(* Logix 5000 project; controller PLC_MCC1201_220AP1 vendor 1 type 14 code 164 rev 35.11; software revision 35.00; part 20 of 25 *)
(* tags used below, declared in another part *)
   LEHR_dActualSpeedValue_mm_min : DINT;
   LEHR_dActualSpeedValueToConveyor_mm_min : DINT;
   LEHR_dLehrPositionAdvancement : DINT;
   SnaprollUPS_DistanceFromSnaproll_cmm : DINT;
   SnaprollUPS_xOS_NewCut : BOOL;
   SnaprollUPS_xOSR : BOOL;
   SnaprollUPS_xOutputRise : BOOL;
   tmOF_retainSnaprolUPS : TIMER;
   TMP_dDummy : DINT;
   TMP_dEncoderCutPosition : DINT;
   TMP_xCutOnSnaproll_cmm : BOOL;
   B3 : DINT[102];
   DISTANCE : ALIAS FOR N7[1];
   M203DROP : MAC_DROPCONV;
   M203DROP_ALM : MAC_DROPCONV_ALM;
   M203DROP_HMR : MAC_DROPCONV_HMR;
   M203DROP_HMW : MAC_DROPCONV_HMW;
   M225 : MAC_EMERGENCYXCUT;
   O : INT[128];
   Status : INT;   // INT tag to retrieve Status value through GSV created during conversion
   TMP_xAlwaysOFF : BOOL;
   TMP_xTestCycle : BOOL;
   W_APC_ACTIVE : ALIAS FOR W_B3[0].10;
   W_APC_BUTTON : ALIAS FOR W_I[8].10;
   W_B3 : DINT[7];
   W_BLOWDOWN_VALVE : ALIAS FOR W_O[10].12;
   W_CB1_START : ALIAS FOR W_O[10].1;
   W_CB2_START : ALIAS FOR W_O[10].3;
   W_COMPUTE_TCD3 : ALIAS FOR W_N7[923];
   W_COMPUTE_TCD5B : ALIAS FOR W_N7[926];
   W_CONDUCT_SENSOR : ALIAS FOR W_N7[110];
   W_CONV_PID_N7_620 : PID;   // Return Water Flow Control Valve Position
   W_CONV_PID_N7_650 : PID;   // RO Unit Water Temperature Control
   W_CONV_PID_N7_680 : PID;   // Boiler Water Temperature Control
   W_CONV_PID_N7_710 : PID;   // Mixed Air Control Damper Positioning
   W_CONV_PID_N7_740 : PID;   // Dryer Room Temperature Control
   W_CP1_ENABLE : ALIAS FOR W_B3[0].5;
   W_CP1A_START : ALIAS FOR W_O[10].5;
   W_CP1B_START : ALIAS FOR W_O[10].7;
   W_CP2A_START : ALIAS FOR W_O[10].9;
   W_CP2B_START : ALIAS FOR W_O[10].11;
   W_DRYER_PID_OUT : ALIAS FOR W_N7[925];
   W_EMER_STOP : ALIAS FOR W_I[8].13;
   W_FLOW_ENABLE : ALIAS FOR W_B3[0].9;
   W_HX1_BCD_OUT : ALIAS FOR W_N7[917];
   W_HX2_SENSOR : ALIAS FOR W_N7[47];
   W_I : INT[32];
   W_MA_FAN_SENSOR : ALIAS FOR W_N7[50];
   W_N11 : DINT[10];
   W_N7 : DINT[933];
   W_PID_INT_TO_TOD : ALIAS FOR W_N7[919];
   W_PS1_SWITCH : ALIAS FOR W_I[8].8;
   W_PWT_HIGH_LIMIT : ALIAS FOR W_I[8].2;
   W_RECIEVING_LEVEL : ALIAS FOR W_I[8].9;
   W_RET_PID_OUTPUT : ALIAS FOR W_N7[921];
   W_RO_START : ALIAS FOR W_O[10].13;
   W_RUN_WASHER : ALIAS FOR W_B3[0].2;
   W_SHUTDOWN_LATCH : ALIAS FOR W_B3[0].1;
   W_T4 : TIMER[101];
   W_TCD3_OUTPUT : ALIAS FOR W_N7[300];
   W_TCD3_PID_OUTPUT : ALIAS FOR W_N7[922];
   W_TCD4_OUTPUT : ALIAS FOR W_N7[301];
   W_TCD5A_OUTPUT : ALIAS FOR W_N7[302];
   W_TT3_RAW_BCD : ALIAS FOR W_N7[48];
   W_TT6_HITEMP_AIR : ALIAS FOR W_N7[49];
   Z200_UPS : ZONE_UPS;
(* MainProgram, continued *)

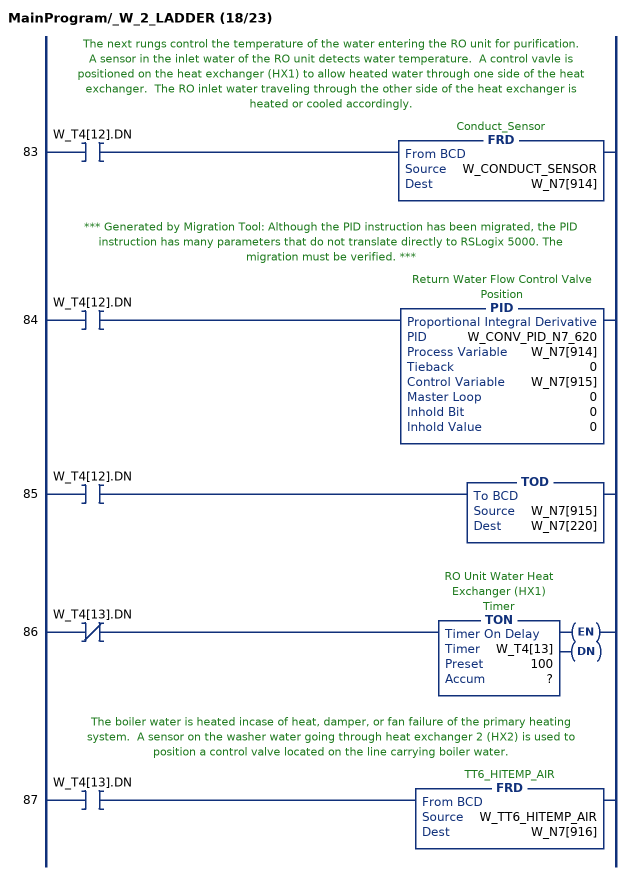
   [picture p330: MainProgram/_W_2_LADDER rungs 83-87]
   // The next rungs control the temperature of the water entering the RO unit for purification.  A sensor in the inlet water of the RO unit detects water temperature.  A control vavle is positioned on the heat exchanger (HX1) to allow heated water through one side of the heat exchanger.  The RO inlet water traveling through the other side of the heat exchanger is heated or cooled accordingly.
   83: XIC(W_T4[12].DN)FRD(W_CONDUCT_SENSOR,W_N7[914]);
   // *** Generated by Migration Tool: Although the PID instruction has been migrated, the PID instruction has many parameters that do not translate directly to RSLogix 5000. The migration must be verified. ***
   84: XIC(W_T4[12].DN)PID(W_CONV_PID_N7_620,W_N7[914],0,W_N7[915],0,0,0);
   85: XIC(W_T4[12].DN)TOD(W_N7[915],W_N7[220]);
   86: XIO(W_T4[13].DN)TON(W_T4[13],?,?);
   // The boiler water is heated incase of heat, damper, or fan failure of the primary heating system.  A sensor on the washer water going through heat exchanger 2 (HX2) is used to position a control valve located on the line carrying boiler water.
   87: XIC(W_T4[13].DN)FRD(W_TT6_HITEMP_AIR,W_N7[916]);
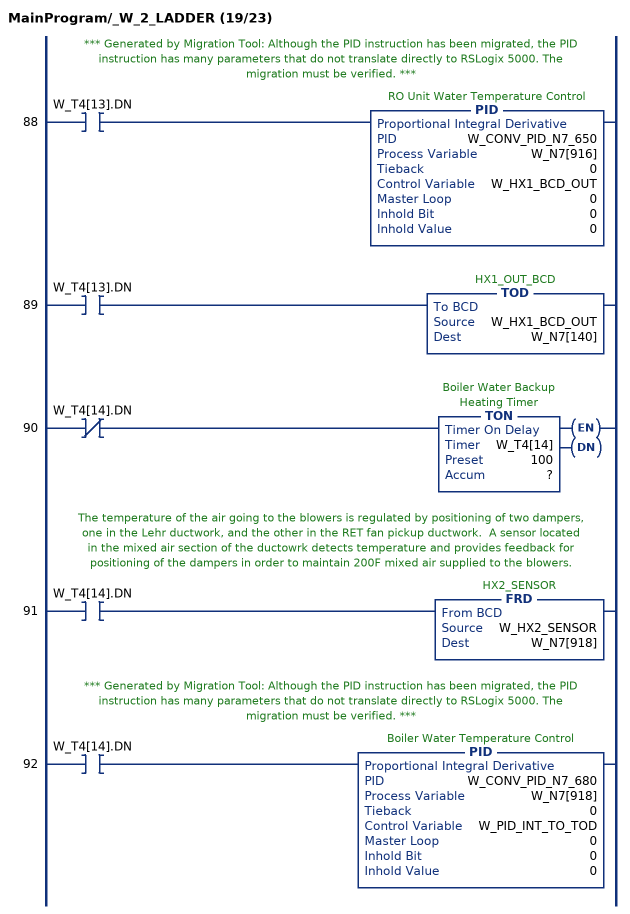
   // *** Generated by Migration Tool: Although the PID instruction has been migrated, the PID instruction has many parameters that do not translate directly to RSLogix 5000. The migration must be verified. ***
   88: XIC(W_T4[13].DN)PID(W_CONV_PID_N7_650,W_N7[916],0,W_HX1_BCD_OUT,0,0,0);
   89: XIC(W_T4[13].DN)TOD(W_HX1_BCD_OUT,W_N7[140]);
   90: XIO(W_T4[14].DN)TON(W_T4[14],?,?);
   // The temperature of the air going to the blowers is regulated by positioning of two dampers, one in the Lehr ductwork, and the other in the RET fan pickup ductwork.  A sensor located in the mixed air section of the ductowrk detects temperature and provides feedback for positioning of the dampers in order to maintain 200F mixed air supplied to the blowers.
   91: XIC(W_T4[14].DN)FRD(W_HX2_SENSOR,W_N7[918]);
   // *** Generated by Migration Tool: Although the PID instruction has been migrated, the PID instruction has many parameters that do not translate directly to RSLogix 5000. The migration must be verified. ***
   92: XIC(W_T4[14].DN)PID(W_CONV_PID_N7_680,W_N7[918],0,W_PID_INT_TO_TOD,0,0,0);
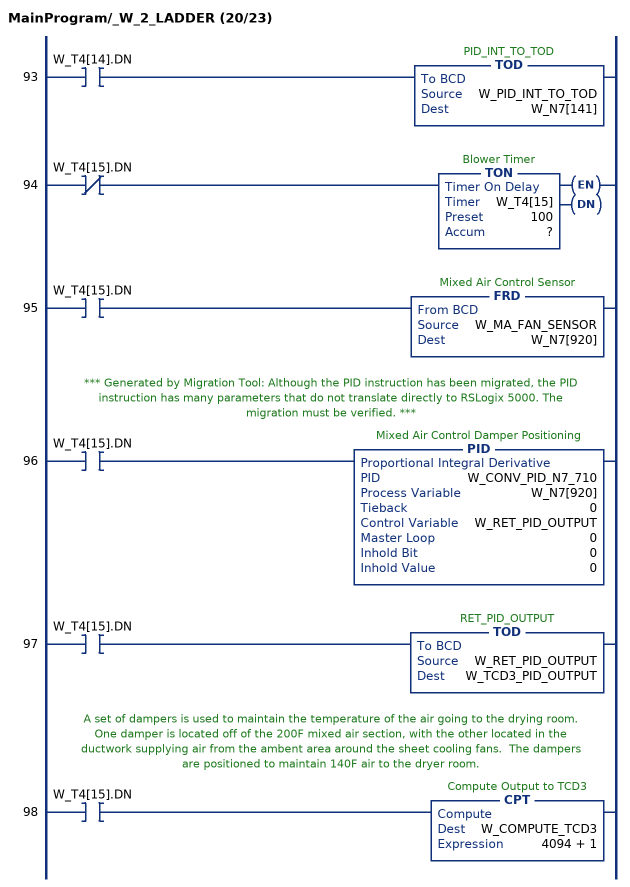
   93: XIC(W_T4[14].DN)TOD(W_PID_INT_TO_TOD,W_N7[141]);
   94: XIO(W_T4[15].DN)TON(W_T4[15],?,?);
   95: XIC(W_T4[15].DN)FRD(W_MA_FAN_SENSOR,W_N7[920]);
   // *** Generated by Migration Tool: Although the PID instruction has been migrated, the PID instruction has many parameters that do not translate directly to RSLogix 5000. The migration must be verified. ***
   96: XIC(W_T4[15].DN)PID(W_CONV_PID_N7_710,W_N7[920],0,W_RET_PID_OUTPUT,0,0,0);
   97: XIC(W_T4[15].DN)TOD(W_RET_PID_OUTPUT,W_TCD3_PID_OUTPUT);
   // A set of dampers is used to maintain the temperature of the air going to the drying room.  One damper is located off of the 200F mixed air section, with the other located in the ductwork supplying air from the ambent area around the sheet cooling fans.  The dampers are positioned to maintain 140F air to the dryer room.
   98: XIC(W_T4[15].DN)CPT(W_COMPUTE_TCD3,4094 + 1);
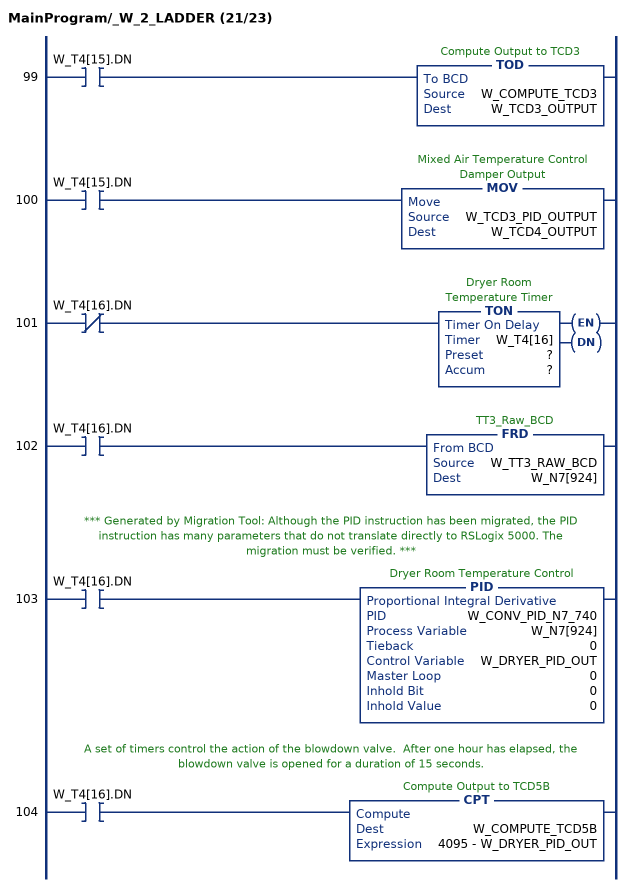
   99: XIC(W_T4[15].DN)TOD(W_COMPUTE_TCD3,W_TCD3_OUTPUT);
   100: XIC(W_T4[15].DN)MOV(W_TCD3_PID_OUTPUT,W_TCD4_OUTPUT);
   101: XIO(W_T4[16].DN)TON(W_T4[16],?,?);
   102: XIC(W_T4[16].DN)FRD(W_TT3_RAW_BCD,W_N7[924]);
   // *** Generated by Migration Tool: Although the PID instruction has been migrated, the PID instruction has many parameters that do not translate directly to RSLogix 5000. The migration must be verified. ***
   103: XIC(W_T4[16].DN)PID(W_CONV_PID_N7_740,W_N7[924],0,W_DRYER_PID_OUT,0,0,0);
   // A set of timers control the action of the blowdown valve.  After one hour has elapsed, the blowdown valve is opened for a duration of 15 seconds.
   104: XIC(W_T4[16].DN)CPT(W_COMPUTE_TCD5B,4095 - W_DRYER_PID_OUT);
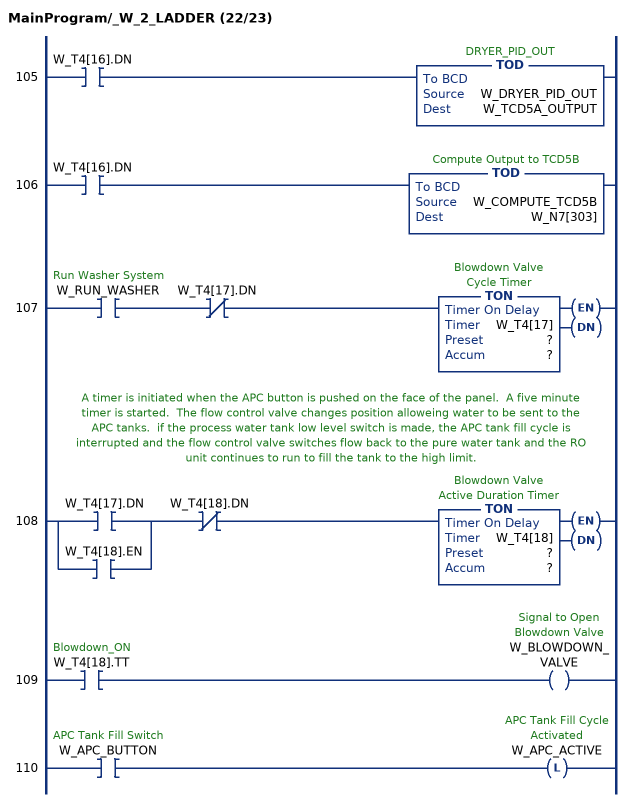
   105: XIC(W_T4[16].DN)TOD(W_DRYER_PID_OUT,W_TCD5A_OUTPUT);
   106: XIC(W_T4[16].DN)TOD(W_COMPUTE_TCD5B,W_N7[303]);
   107: XIC(W_RUN_WASHER)XIO(W_T4[17].DN)TON(W_T4[17],?,?);
   // A timer is initiated when the APC button is pushed on the face of the panel.  A five minute timer is started.  The flow control valve changes position alloweing water to be sent to the APC tanks.  if the process water tank low level switch is made, the APC tank fill cycle is interrupted and the flow control valve switches flow back to the pure water tank and the RO unit continues to run to fill the tank to the high limit.
   108: [XIC(W_T4[17].DN) ,XIC(W_T4[18].EN) ]XIO(W_T4[18].DN)TON(W_T4[18],?,?);
   109: XIC(W_T4[18].TT)OTE(W_BLOWDOWN_VALVE);
   110: XIC(W_APC_BUTTON)OTL(W_APC_ACTIVE);
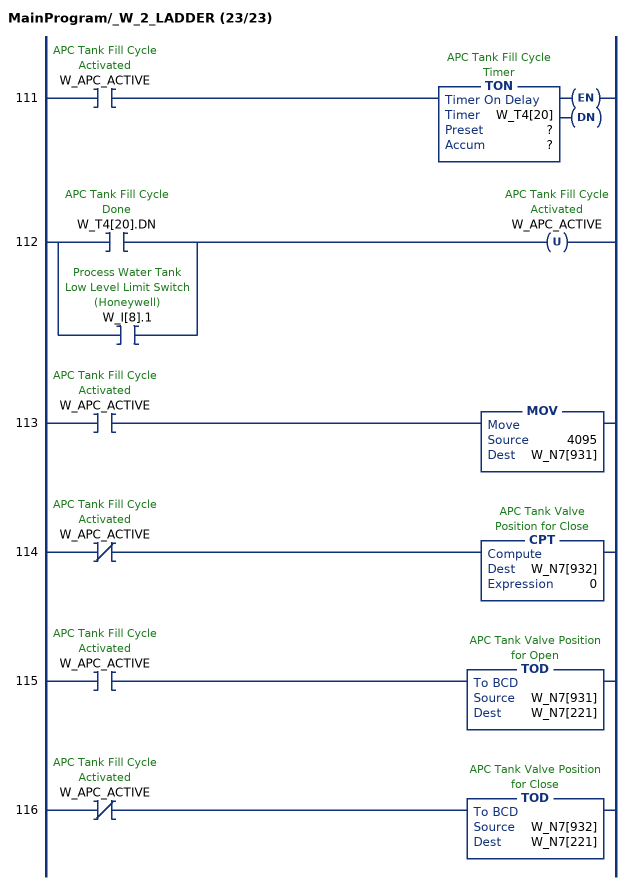
   111: XIC(W_APC_ACTIVE)TON(W_T4[20],?,?);
   112: [XIC(W_T4[20].DN) ,XIC(W_I[8].1) ]OTU(W_APC_ACTIVE);
   113: XIC(W_APC_ACTIVE)MOV(4095,W_N7[931]);
   114: XIO(W_APC_ACTIVE)CPT(W_N7[932],0);
   115: XIC(W_APC_ACTIVE)TOD(W_N7[931],W_N7[221]);
   116: XIO(W_APC_ACTIVE)TOD(W_N7[932],W_N7[221]);
END_ROUTINE

ROUTINE _W_5_LADDER   (* ladder *)
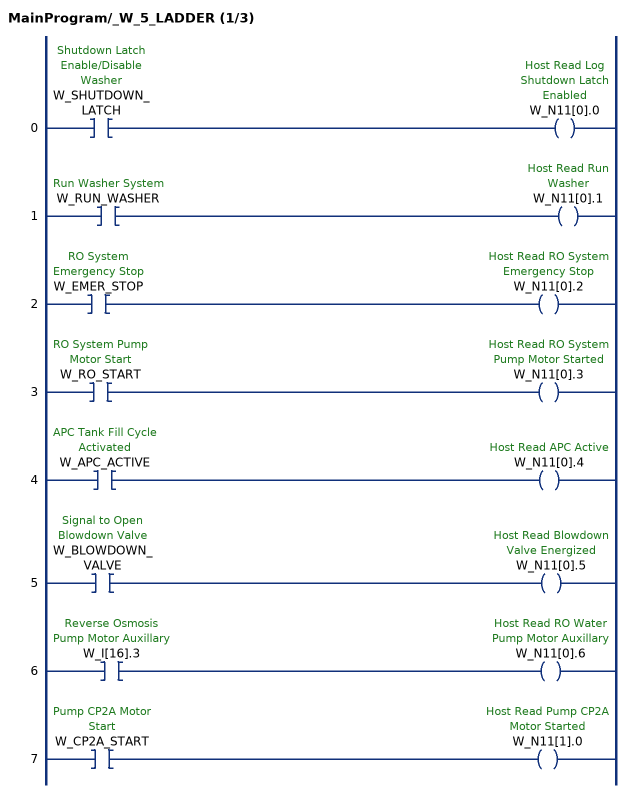
   0: XIC(W_SHUTDOWN_LATCH)OTE(W_N11[0].0);
   1: XIC(W_RUN_WASHER)OTE(W_N11[0].1);
   2: XIC(W_EMER_STOP)OTE(W_N11[0].2);
   3: XIC(W_RO_START)OTE(W_N11[0].3);
   4: XIC(W_APC_ACTIVE)OTE(W_N11[0].4);
   5: XIC(W_BLOWDOWN_VALVE)OTE(W_N11[0].5);
   6: XIC(W_I[16].3)OTE(W_N11[0].6);
   7: XIC(W_CP2A_START)OTE(W_N11[1].0);
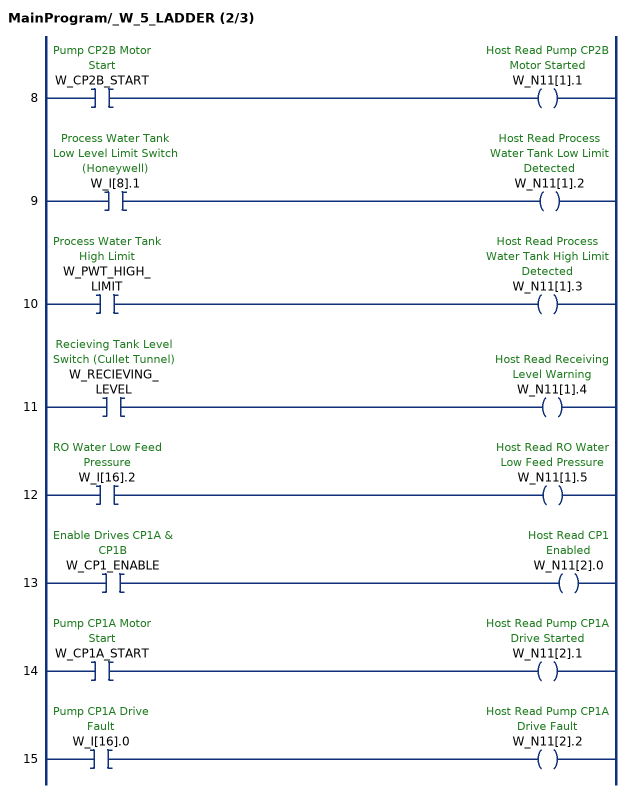
   8: XIC(W_CP2B_START)OTE(W_N11[1].1);
   9: XIC(W_I[8].1)OTE(W_N11[1].2);
   10: XIC(W_PWT_HIGH_LIMIT)OTE(W_N11[1].3);
   11: XIC(W_RECIEVING_LEVEL)OTE(W_N11[1].4);
   12: XIC(W_I[16].2)OTE(W_N11[1].5);
   13: XIC(W_CP1_ENABLE)OTE(W_N11[2].0);
   14: XIC(W_CP1A_START)OTE(W_N11[2].1);
   15: XIC(W_I[16].0)OTE(W_N11[2].2);
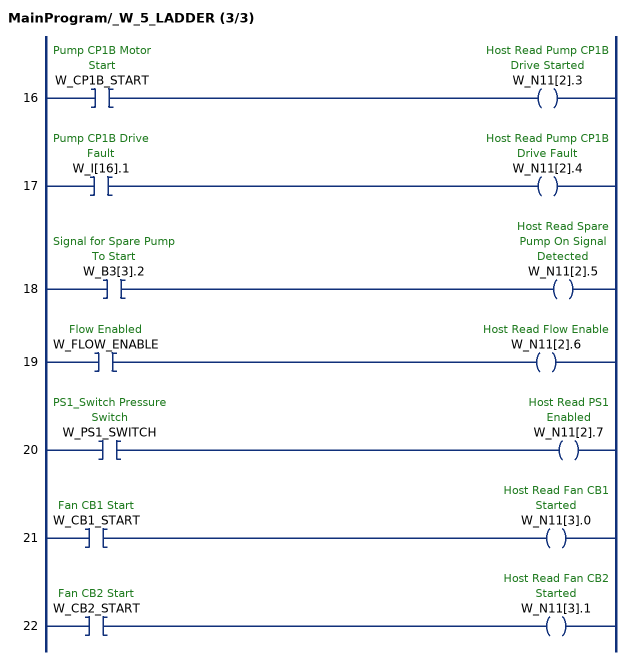
   16: XIC(W_CP1B_START)OTE(W_N11[2].3);
   17: XIC(W_I[16].1)OTE(W_N11[2].4);
   18: XIC(W_B3[3].2)OTE(W_N11[2].5);
   19: XIC(W_FLOW_ENABLE)OTE(W_N11[2].6);
   20: XIC(W_PS1_SWITCH)OTE(W_N11[2].7);
   21: XIC(W_CB1_START)OTE(W_N11[3].0);
   22: XIC(W_CB2_START)OTE(W_N11[3].1);
END_ROUTINE

ROUTINE Conveyors_Logic   (* ladder *)
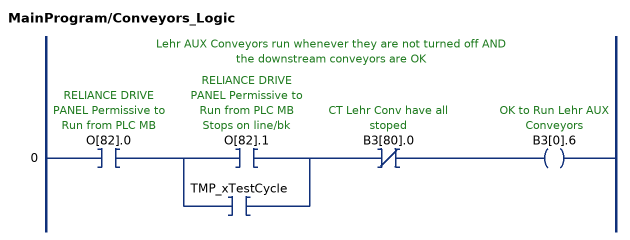
   // Lehr AUX Conveyors run whenever they are not turned off AND
   // the downstream conveyors are OK
   0: XIC(O[82].0)[XIC(O[82].1) ,XIC(TMP_xTestCycle) ]XIO(B3[80].0)OTE(B3[0].6);
END_ROUTINE

ROUTINE M203_DropConveyor_Faults   (* ladder *)
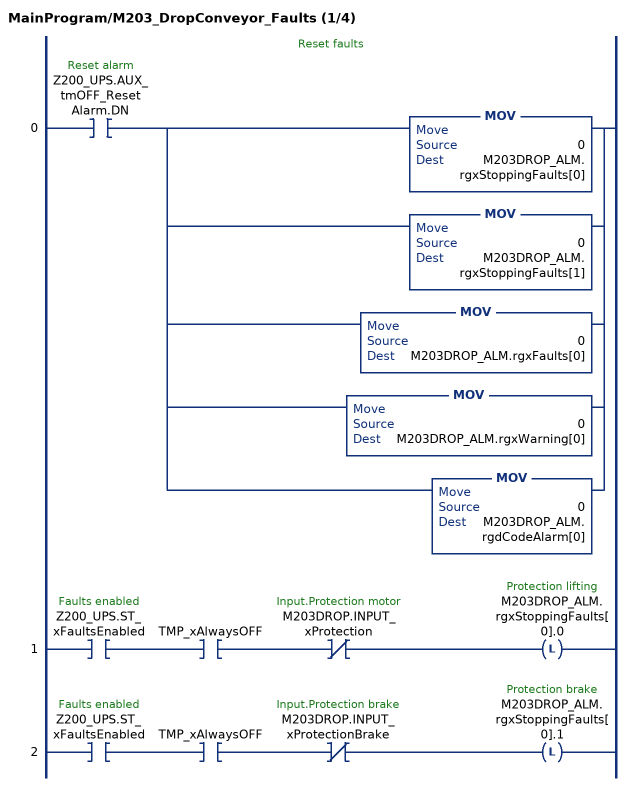
   // Reset faults
   0: XIC(Z200_UPS.AUX_tmOFF_ResetAlarm.DN)[MOV(0,M203DROP_ALM.rgxStoppingFaults[0]) ,MOV(0,M203DROP_ALM.rgxStoppingFaults[1]) ,MOV(0,M203DROP_ALM.rgxFaults[0]) ,MOV(0,M203DROP_ALM.rgxWarning[0]) ,MOV(0,M203DROP_ALM.rgdCodeAlarm[0]) ];
   1: XIC(Z200_UPS.ST_xFaultsEnabled)XIC(TMP_xAlwaysOFF)XIO(M203DROP.INPUT_xProtection)OTL(M203DROP_ALM.rgxStoppingFaults[0].0);
   2: XIC(Z200_UPS.ST_xFaultsEnabled)XIC(TMP_xAlwaysOFF)XIO(M203DROP.INPUT_xProtectionBrake)OTL(M203DROP_ALM.rgxStoppingFaults[0].1);
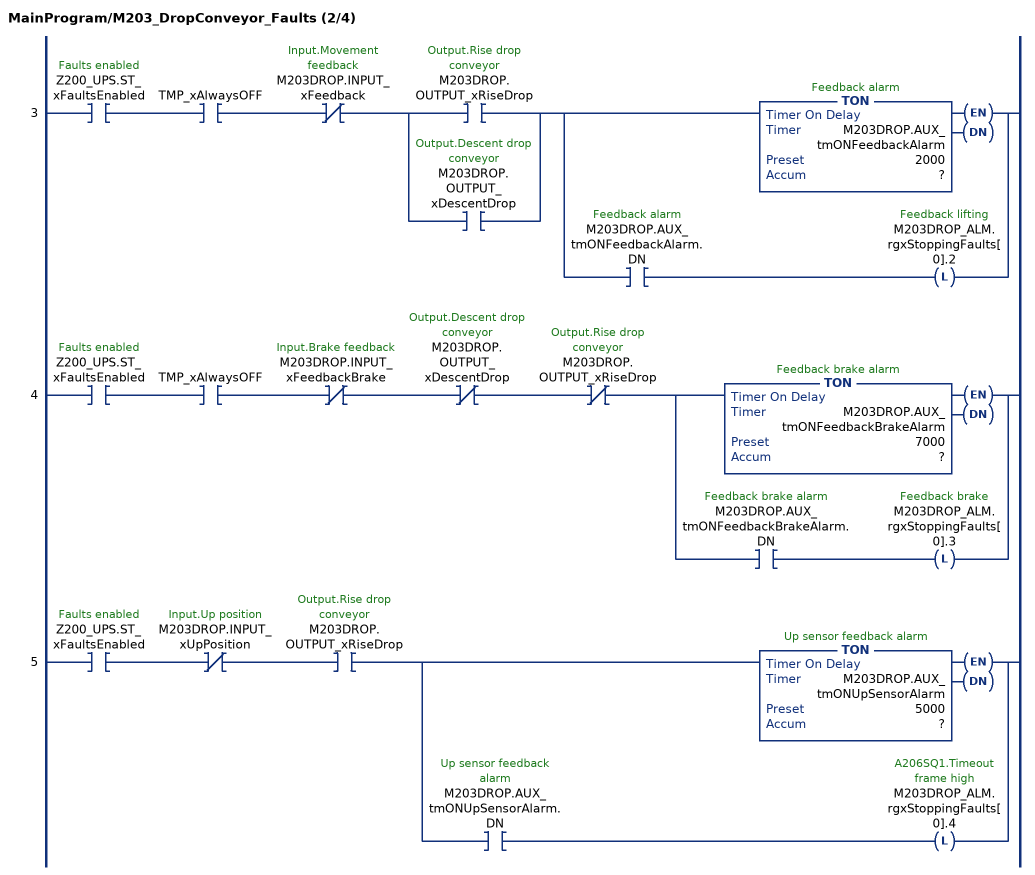
   3: XIC(Z200_UPS.ST_xFaultsEnabled)XIC(TMP_xAlwaysOFF)XIO(M203DROP.INPUT_xFeedback)[XIC(M203DROP.OUTPUT_xRiseDrop) ,XIC(M203DROP.OUTPUT_xDescentDrop) ][TON(M203DROP.AUX_tmONFeedbackAlarm,?,?) ,XIC(M203DROP.AUX_tmONFeedbackAlarm.DN) OTL(M203DROP_ALM.rgxStoppingFaults[0].2) ];
   4: XIC(Z200_UPS.ST_xFaultsEnabled)XIC(TMP_xAlwaysOFF)XIO(M203DROP.INPUT_xFeedbackBrake)XIO(M203DROP.OUTPUT_xDescentDrop)XIO(M203DROP.OUTPUT_xRiseDrop)[TON(M203DROP.AUX_tmONFeedbackBrakeAlarm,?,?) ,XIC(M203DROP.AUX_tmONFeedbackBrakeAlarm.DN) OTL(M203DROP_ALM.rgxStoppingFaults[0].3) ];
   5: XIC(Z200_UPS.ST_xFaultsEnabled)XIO(M203DROP.INPUT_xUpPosition)XIC(M203DROP.OUTPUT_xRiseDrop)[TON(M203DROP.AUX_tmONUpSensorAlarm,?,?) ,XIC(M203DROP.AUX_tmONUpSensorAlarm.DN) OTL(M203DROP_ALM.rgxStoppingFaults[0].4) ];
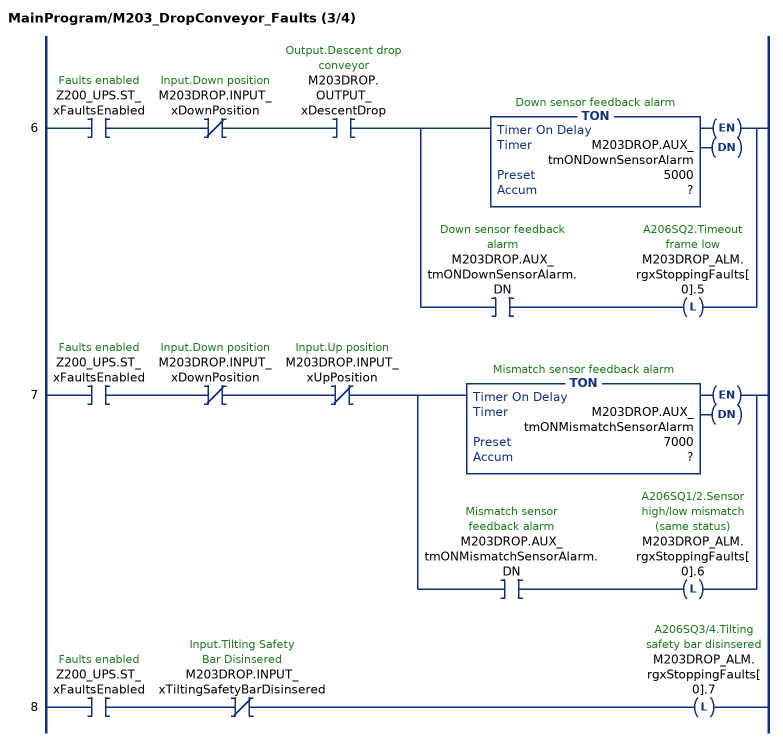
   6: XIC(Z200_UPS.ST_xFaultsEnabled)XIO(M203DROP.INPUT_xDownPosition)XIC(M203DROP.OUTPUT_xDescentDrop)[TON(M203DROP.AUX_tmONDownSensorAlarm,?,?) ,XIC(M203DROP.AUX_tmONDownSensorAlarm.DN) OTL(M203DROP_ALM.rgxStoppingFaults[0].5) ];
   7: XIC(Z200_UPS.ST_xFaultsEnabled)XIO(M203DROP.INPUT_xDownPosition)XIO(M203DROP.INPUT_xUpPosition)[TON(M203DROP.AUX_tmONMismatchSensorAlarm,?,?) ,XIC(M203DROP.AUX_tmONMismatchSensorAlarm.DN) OTL(M203DROP_ALM.rgxStoppingFaults[0].6) ];
   8: XIC(Z200_UPS.ST_xFaultsEnabled)XIO(M203DROP.INPUT_xTiltingSafetyBarDisinsered)OTL(M203DROP_ALM.rgxStoppingFaults[0].7);
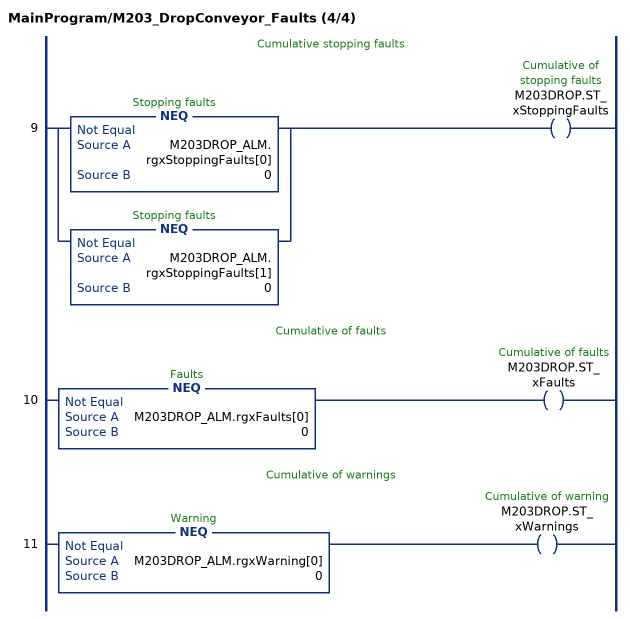
   // Cumulative stopping faults
   9: [NEQ(M203DROP_ALM.rgxStoppingFaults[0],0) ,NEQ(M203DROP_ALM.rgxStoppingFaults[1],0) ]OTE(M203DROP.ST_xStoppingFaults);
   // Cumulative of faults
   10: NEQ(M203DROP_ALM.rgxFaults[0],0)OTE(M203DROP.ST_xFaults);
   // Cumulative of warnings
   11: NEQ(M203DROP_ALM.rgxWarning[0],0)OTE(M203DROP.ST_xWarnings);
END_ROUTINE

ROUTINE M203_DropConveyor_Logics   (* ladder *)
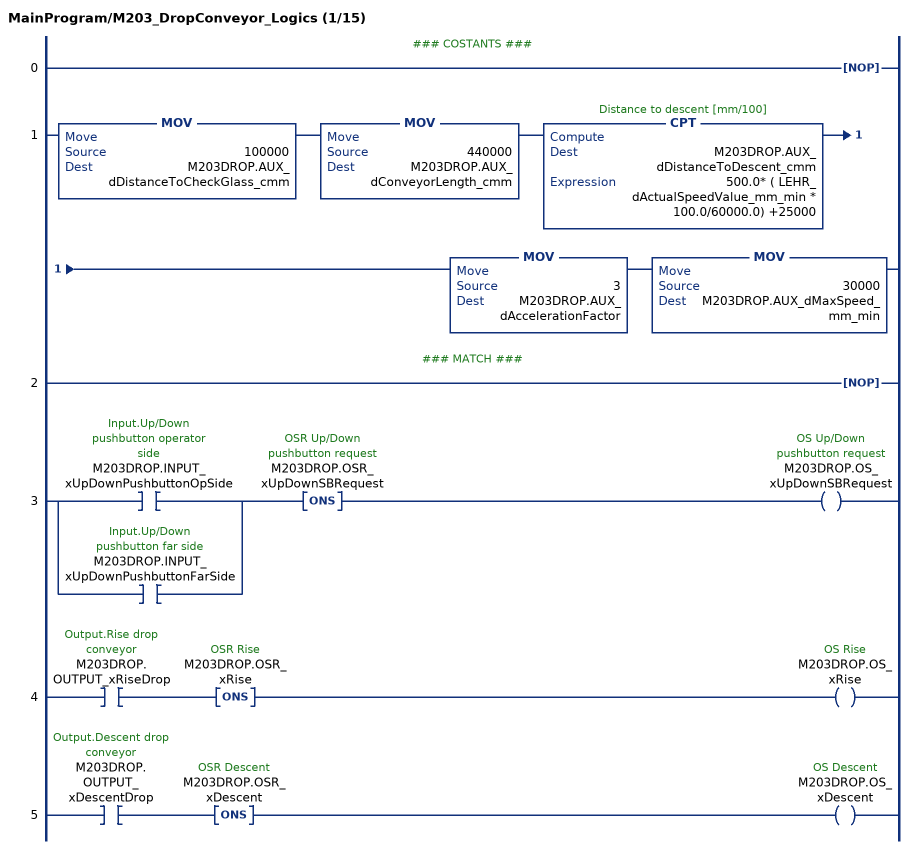
   // ### COSTANTS ###
   0: NOP();
   1: MOV(100000,M203DROP.AUX_dDistanceToCheckGlass_cmm)MOV(440000,M203DROP.AUX_dConveyorLength_cmm)CPT(M203DROP.AUX_dDistanceToDescent_cmm,500.0* ( LEHR_dActualSpeedValue_mm_min * 100.0/60000.0) +25000)MOV(3,M203DROP.AUX_dAccelerationFactor)MOV(30000,M203DROP.AUX_dMaxSpeed_mm_min);
   // ### MATCH ###
   2: NOP();
   3: [XIC(M203DROP.INPUT_xUpDownPushbuttonOpSide) ,XIC(M203DROP.INPUT_xUpDownPushbuttonFarSide) ]ONS(M203DROP.OSR_xUpDownSBRequest)OTE(M203DROP.OS_xUpDownSBRequest);
   4: XIC(M203DROP.OUTPUT_xRiseDrop)ONS(M203DROP.OSR_xRise)OTE(M203DROP.OS_xRise);
   5: XIC(M203DROP.OUTPUT_xDescentDrop)ONS(M203DROP.OSR_xDescent)OTE(M203DROP.OS_xDescent);
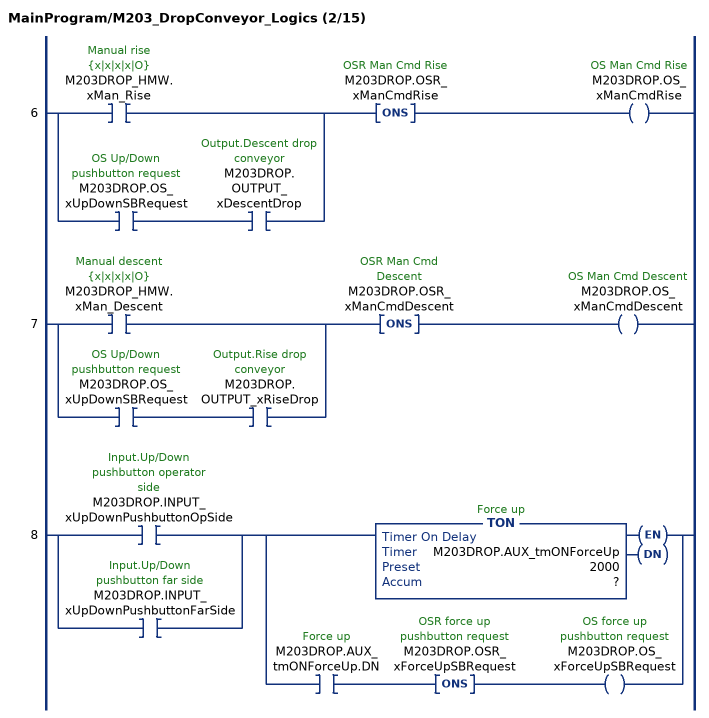
   6: [XIC(M203DROP_HMW.xMan_Rise) ,XIC(M203DROP.OS_xUpDownSBRequest) XIC(M203DROP.OUTPUT_xDescentDrop) ]ONS(M203DROP.OSR_xManCmdRise)OTE(M203DROP.OS_xManCmdRise);
   7: [XIC(M203DROP_HMW.xMan_Descent) ,XIC(M203DROP.OS_xUpDownSBRequest) XIC(M203DROP.OUTPUT_xRiseDrop) ]ONS(M203DROP.OSR_xManCmdDescent)OTE(M203DROP.OS_xManCmdDescent);
   8: [XIC(M203DROP.INPUT_xUpDownPushbuttonOpSide) ,XIC(M203DROP.INPUT_xUpDownPushbuttonFarSide) ][TON(M203DROP.AUX_tmONForceUp,?,?) ,XIC(M203DROP.AUX_tmONForceUp.DN) ONS(M203DROP.OSR_xForceUpSBRequest) OTE(M203DROP.OS_xForceUpSBRequest) ];
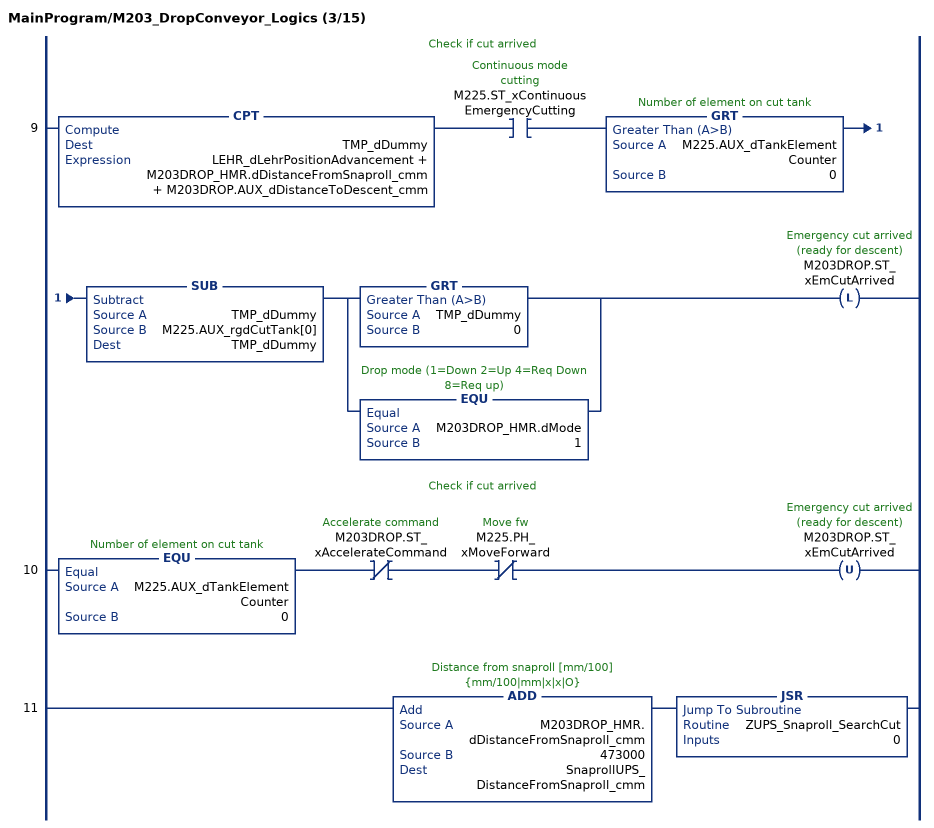
   // Check if cut arrived
   9: CPT(TMP_dDummy,LEHR_dLehrPositionAdvancement + M203DROP_HMR.dDistanceFromSnaproll_cmm + M203DROP.AUX_dDistanceToDescent_cmm)XIC(M225.ST_xContinuousEmergencyCutting)GRT(M225.AUX_dTankElementCounter,0)SUB(TMP_dDummy,M225.AUX_rgdCutTank[0],TMP_dDummy)[GRT(TMP_dDummy,0) ,EQU(M203DROP_HMR.dMode,1) ]OTL(M203DROP.ST_xEmCutArrived);
   // Check if cut arrived
   10: EQU(M225.AUX_dTankElementCounter,0)XIO(M203DROP.ST_xAccelerateCommand)XIO(M225.PH_xMoveForward)OTU(M203DROP.ST_xEmCutArrived);
   11: ADD(M203DROP_HMR.dDistanceFromSnaproll_cmm,473000,SnaprollUPS_DistanceFromSnaproll_cmm)JSR(ZUPS_Snaproll_SearchCut,0);
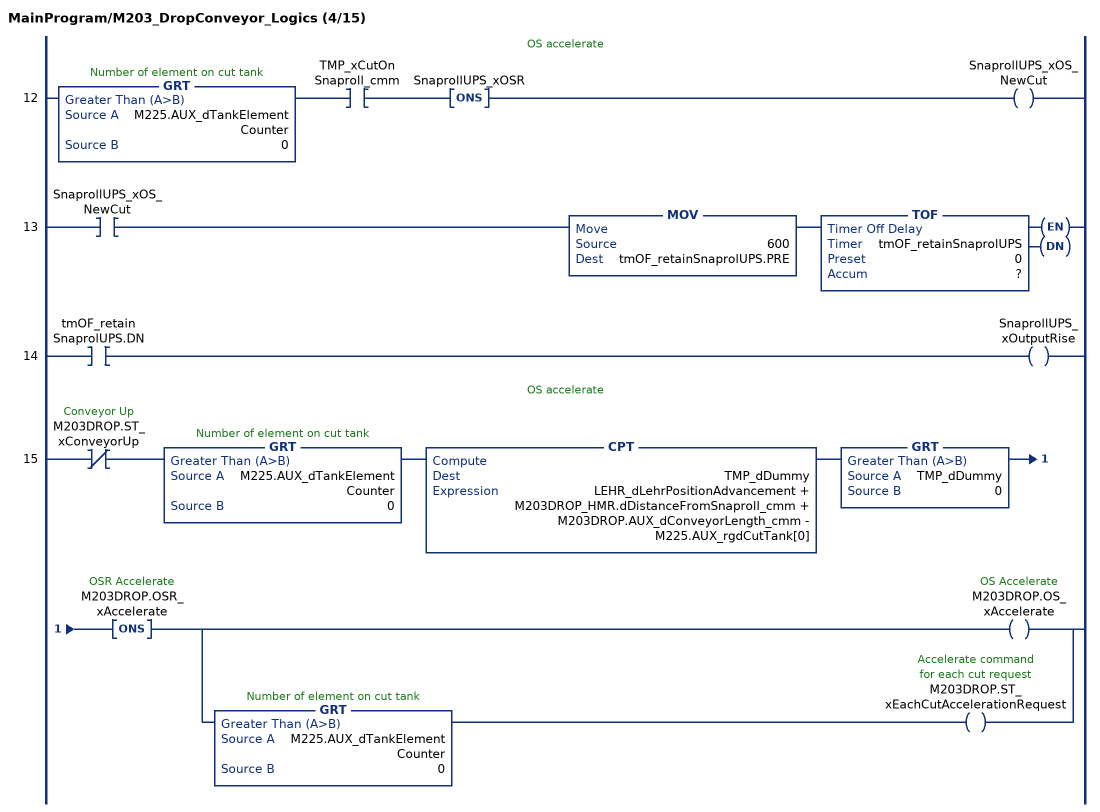
   // OS accelerate
   12: GRT(M225.AUX_dTankElementCounter,0)XIC(TMP_xCutOnSnaproll_cmm)ONS(SnaprollUPS_xOSR)OTE(SnaprollUPS_xOS_NewCut);
   13: XIC(SnaprollUPS_xOS_NewCut)MOV(600,tmOF_retainSnaprolUPS.PRE)TOF(tmOF_retainSnaprolUPS,?,?);
   14: XIC(tmOF_retainSnaprolUPS.DN)OTE(SnaprollUPS_xOutputRise);
   // OS accelerate
   15: XIO(M203DROP.ST_xConveyorUp)GRT(M225.AUX_dTankElementCounter,0)CPT(TMP_dDummy,LEHR_dLehrPositionAdvancement + M203DROP_HMR.dDistanceFromSnaproll_cmm + M203DROP.AUX_dConveyorLength_cmm - M225.AUX_rgdCutTank[0])GRT(TMP_dDummy,0)ONS(M203DROP.OSR_xAccelerate)[OTE(M203DROP.OS_xAccelerate) ,GRT(M225.AUX_dTankElementCounter,0) OTE(M203DROP.ST_xEachCutAccelerationRequest) ];
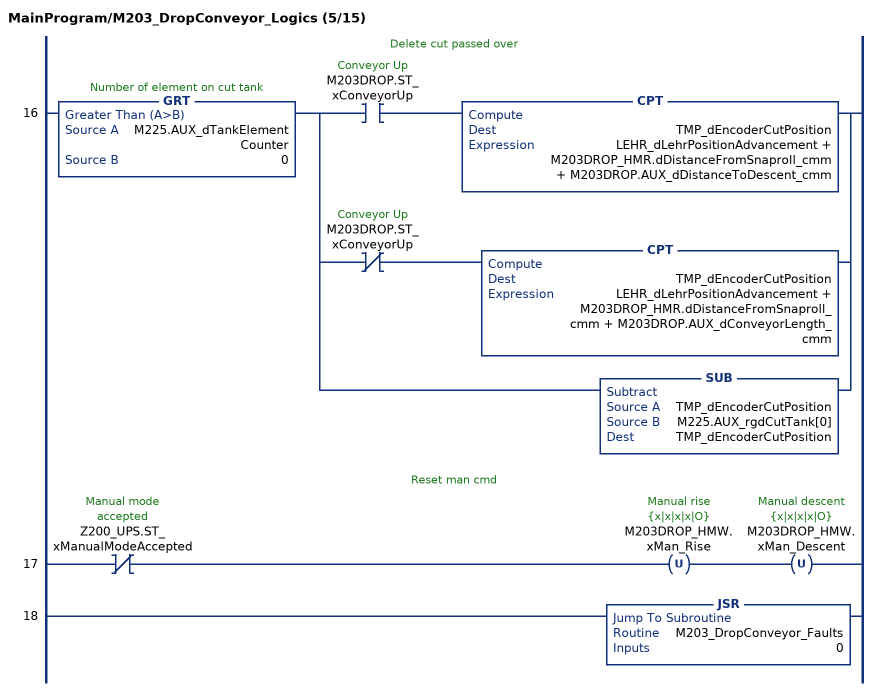
   // Delete cut passed over
   16: GRT(M225.AUX_dTankElementCounter,0)[XIC(M203DROP.ST_xConveyorUp) CPT(TMP_dEncoderCutPosition,LEHR_dLehrPositionAdvancement + M203DROP_HMR.dDistanceFromSnaproll_cmm + M203DROP.AUX_dDistanceToDescent_cmm) ,XIO(M203DROP.ST_xConveyorUp) CPT(TMP_dEncoderCutPosition,LEHR_dLehrPositionAdvancement + M203DROP_HMR.dDistanceFromSnaproll_cmm + M203DROP.AUX_dConveyorLength_cmm) ,SUB(TMP_dEncoderCutPosition,M225.AUX_rgdCutTank[0],TMP_dEncoderCutPosition) ];
   // Reset man cmd
   17: XIO(Z200_UPS.ST_xManualModeAccepted)OTU(M203DROP_HMW.xMan_Rise)OTU(M203DROP_HMW.xMan_Descent);
   18: JSR(M203_DropConveyor_Faults,0);
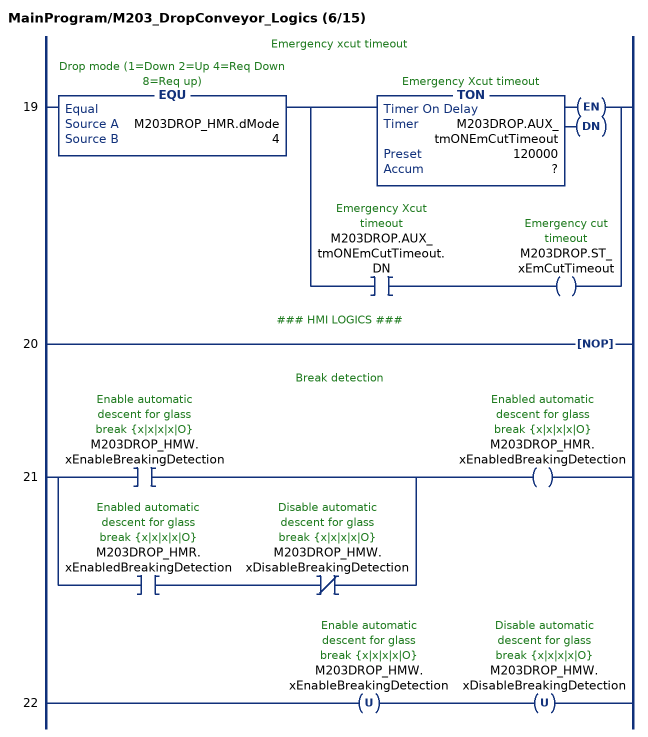
   // Emergency xcut timeout
   19: EQU(M203DROP_HMR.dMode,4)[TON(M203DROP.AUX_tmONEmCutTimeout,?,?) ,XIC(M203DROP.AUX_tmONEmCutTimeout.DN) OTE(M203DROP.ST_xEmCutTimeout) ];
   // ### HMI LOGICS ###
   20: NOP();
   // Break detection
   21: [XIC(M203DROP_HMW.xEnableBreakingDetection) ,XIC(M203DROP_HMR.xEnabledBreakingDetection) XIO(M203DROP_HMW.xDisableBreakingDetection) ]OTE(M203DROP_HMR.xEnabledBreakingDetection);
   22: OTU(M203DROP_HMW.xEnableBreakingDetection)OTU(M203DROP_HMW.xDisableBreakingDetection);
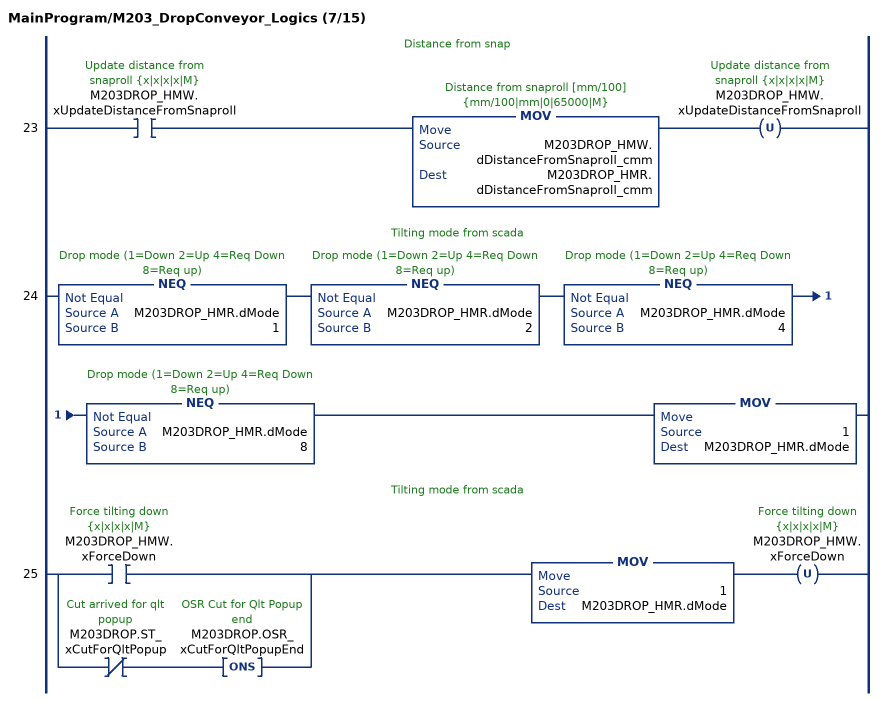
   // Distance from snap
   23: XIC(M203DROP_HMW.xUpdateDistanceFromSnaproll)MOV(M203DROP_HMW.dDistanceFromSnaproll_cmm,M203DROP_HMR.dDistanceFromSnaproll_cmm)OTU(M203DROP_HMW.xUpdateDistanceFromSnaproll);
   // Tilting mode from scada
   24: NEQ(M203DROP_HMR.dMode,1)NEQ(M203DROP_HMR.dMode,2)NEQ(M203DROP_HMR.dMode,4)NEQ(M203DROP_HMR.dMode,8)MOV(1,M203DROP_HMR.dMode);
   // Tilting mode from scada
   25: [XIC(M203DROP_HMW.xForceDown) ,XIO(M203DROP.ST_xCutForQltPopup) ONS(M203DROP.OSR_xCutForQltPopupEnd) ]MOV(1,M203DROP_HMR.dMode)OTU(M203DROP_HMW.xForceDown);
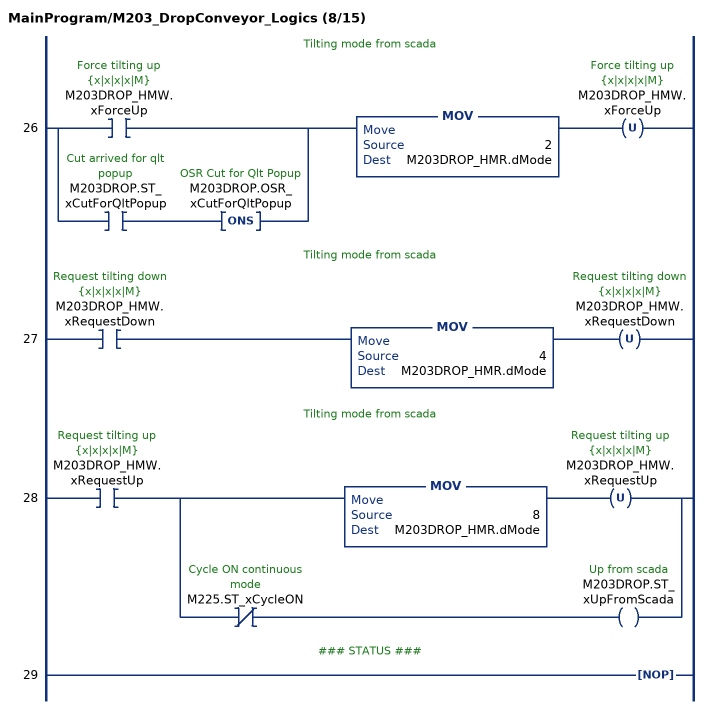
   // Tilting mode from scada
   26: [XIC(M203DROP_HMW.xForceUp) ,XIC(M203DROP.ST_xCutForQltPopup) ONS(M203DROP.OSR_xCutForQltPopup) ]MOV(2,M203DROP_HMR.dMode)OTU(M203DROP_HMW.xForceUp);
   // Tilting mode from scada
   27: XIC(M203DROP_HMW.xRequestDown)MOV(4,M203DROP_HMR.dMode)OTU(M203DROP_HMW.xRequestDown);
   // Tilting mode from scada
   28: XIC(M203DROP_HMW.xRequestUp)[MOV(8,M203DROP_HMR.dMode) OTU(M203DROP_HMW.xRequestUp) ,XIO(M225.ST_xCycleON) OTE(M203DROP.ST_xUpFromScada) ];
   // ### STATUS ###
   29: NOP();
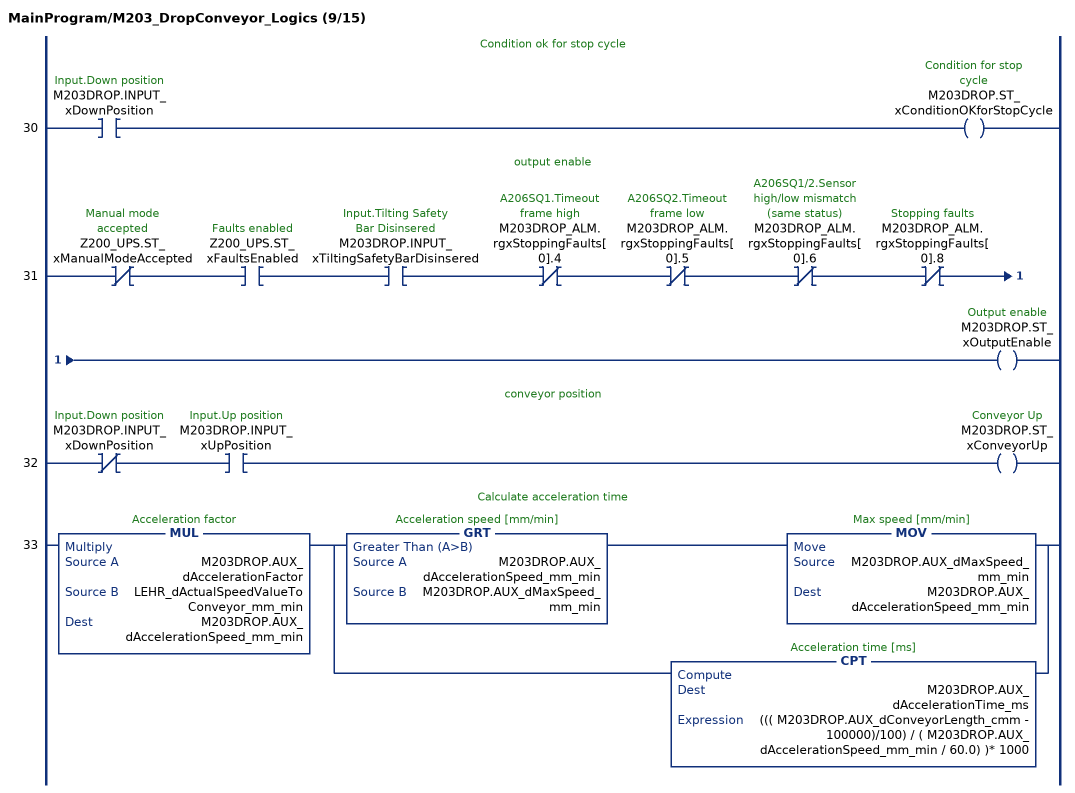
   // Condition ok for stop cycle
   30: XIC(M203DROP.INPUT_xDownPosition)OTE(M203DROP.ST_xConditionOKforStopCycle);
   // output enable
   31: XIO(Z200_UPS.ST_xManualModeAccepted)XIC(Z200_UPS.ST_xFaultsEnabled)XIC(M203DROP.INPUT_xTiltingSafetyBarDisinsered)XIO(M203DROP_ALM.rgxStoppingFaults[0].4)XIO(M203DROP_ALM.rgxStoppingFaults[0].5)XIO(M203DROP_ALM.rgxStoppingFaults[0].6)XIO(M203DROP_ALM.rgxStoppingFaults[0].8)OTE(M203DROP.ST_xOutputEnable);
   // conveyor position
   32: XIO(M203DROP.INPUT_xDownPosition)XIC(M203DROP.INPUT_xUpPosition)OTE(M203DROP.ST_xConveyorUp);
   // Calculate acceleration time
   33: MUL(M203DROP.AUX_dAccelerationFactor,LEHR_dActualSpeedValueToConveyor_mm_min,M203DROP.AUX_dAccelerationSpeed_mm_min)[GRT(M203DROP.AUX_dAccelerationSpeed_mm_min,M203DROP.AUX_dMaxSpeed_mm_min) MOV(M203DROP.AUX_dMaxSpeed_mm_min,M203DROP.AUX_dAccelerationSpeed_mm_min) ,CPT(M203DROP.AUX_dAccelerationTime_ms,((( M203DROP.AUX_dConveyorLength_cmm - 100000)/100) / ( M203DROP.AUX_dAccelerationSpeed_mm_min / 60.0) )* 1000) ];
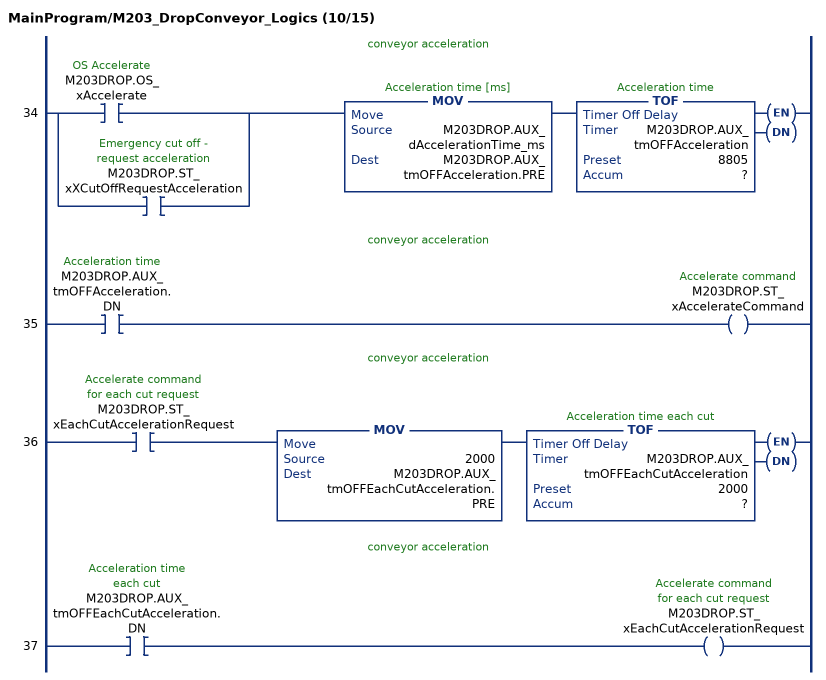
   // conveyor acceleration
   34: [XIC(M203DROP.OS_xAccelerate) ,XIC(M203DROP.ST_xXCutOffRequestAcceleration) ]MOV(M203DROP.AUX_dAccelerationTime_ms,M203DROP.AUX_tmOFFAcceleration.PRE)TOF(M203DROP.AUX_tmOFFAcceleration,?,?);
   // conveyor acceleration
   35: XIC(M203DROP.AUX_tmOFFAcceleration.DN)OTE(M203DROP.ST_xAccelerateCommand);
   // conveyor acceleration
   36: XIC(M203DROP.ST_xEachCutAccelerationRequest)MOV(2000,M203DROP.AUX_tmOFFEachCutAcceleration.PRE)TOF(M203DROP.AUX_tmOFFEachCutAcceleration,?,?);
   // conveyor acceleration
   37: XIC(M203DROP.AUX_tmOFFEachCutAcceleration.DN)OTE(M203DROP.ST_xEachCutAccelerationRequest);
